   "Carrier_40_G120DStatusWord.3" AT %I2362.3 : Bool;   // Bit_03_FAULT
   "Carrier_40_G120DStatusWord.4" AT %I2362.4 : Bool;   // Bit_04_OFF2
   "Carrier_40_G120DStatusWord.5" AT %I2362.5 : Bool;   // Bit_05_OFF3
   "Carrier_40_G120DStatusWord.6" AT %I2362.6 : Bool;   // Bit_06_LOCK_OUT
   "Carrier_40_G120DStatusWord.7" AT %I2362.7 : Bool;   // Bit_07_WARN
   "Carrier_40_G120DStatusWord.8" AT %I2363.0 : Bool;   // Bit_08_NO_DEVIATION
   "Carrier_40_G120DStatusWord.9" AT %I2363.1 : Bool;   // Bit_09_CONTR_PLC
   "Carrier_40_G120DStatusWord.10" AT %I2363.2 : Bool;   // Bit_10_F_MAX
   "Carrier_40_G120DStatusWord.11" AT %I2363.3 : Bool;   // Bit_11_LIMIT_REACHED
   "Carrier_40_G120DStatusWord.12" AT %I2363.4 : Bool;   // Bit_12_BRAKE_OPEN
   "Carrier_40_G120DStatusWord.13" AT %I2363.5 : Bool;   // Bit_13_NO_OVERTEMP
   "Carrier_40_G120DStatusWord.14" AT %I2363.6 : Bool;   // Bit_14_CW_CCW
   "Carrier_40_G120DStatusWord.15" AT %I2363.7 : Bool;   // Bit_15_OVERL
   "Carrier_40_Slot2_Input" AT %IW2364 : Word;   // SLOT 2 INPUT WORD
   "Carrier_40_CrashDetectSW" AT %I2364.0 : Bool;   // CRASH DETECT SW
   "Carrier_40_SpareSafetyInput(2_1)" AT %I2364.1 : Bool;   // SPARE SAFETY INPUT
   "Carrier_40_SpareSafetyInput(2_2)" AT %I2364.2 : Bool;   // SPARE SAFETY INPUT
   "Carrier_40_SpareSafetyInput(2_3)" AT %I2364.3 : Bool;   // SPARE SAFETY INPUT
   "Carrier_40_SpareSafetyInput(2_4)" AT %I2364.4 : Bool;   // SPARE SAFETY INPUT
   "Carrier_40_SpareSafetyInput(2_5)" AT %I2364.5 : Bool;   // SPARE SAFETY INPUT
   "Carrier_40_SpareSafetyInput(2_6)" AT %I2364.6 : Bool;   // SPARE SAFETY INPUT
   "Carrier_40_SpareSafetyInput(2_7)" AT %I2364.7 : Bool;   // SPARE SAFETY INPUT
   "Carrier_40_Slot3_SafetyOutput" AT %IW2365 : Word;   // SLOT 3 SAFETY OUTPUT WORD
   "Carrier_40_Crash_Detect_OK" AT %I2365.0 : Bool;   // CARRIER CRASH DETECT
   "Carrier_40_SpareSafetyOutput(3_1)" AT %I2365.1 : Bool;   // SPARE SAFETY OUTPUT
   "Carrier_40_SpareSafetyOutput(3_2)" AT %I2365.2 : Bool;   // SPARE SAFETY OUTPUT
   "Carrier_40_SpareSafetyOutput(3_3)" AT %I2365.3 : Bool;   // SPARE SAFETY OUTPUT
   "Carrier_40_SpareSafetyOutput(3_4)" AT %I2365.4 : Bool;   // SPARE SAFETY OUTPUT
   "Carrier_40_SpareSafetyOutput(3_5)" AT %I2365.5 : Bool;   // SPARE SAFETY OUTPUT
   "Carrier_40_SpareSafetyOutput(3_6)" AT %I2365.6 : Bool;   // SPARE SAFETY OUTPUT
   "Carrier_40_SpareSafetyOutput(3_7)" AT %I2365.7 : Bool;   // SPARE SAFETY OUTPUT
   "Carrier_40_Slot4_Input" AT %IW2366 : Word;   // SLOT 4 INPUT WORD
   "Carrier_40_480VPowerOn_MDCB1" AT %I2366.0 : Bool;   // 480 VAC POWER ON MDCB 1
   "Carrier_40_SpareInput(4_1)" AT %I2366.1 : Bool;   // SPARE INPUT
   "Carrier_40_SpareInput(4_2)" AT %I2366.2 : Bool;   // SPARE INPUT
   "Carrier_40_SitopSelectStatus" AT %I2366.3 : Bool;   // SITOP SELECT STATUS
   "Carrier_40_DCsupplyOnPSCB2" AT %I2366.4 : Bool;   // DC SUPPLY ON PSCB 2
   "Carrier_40_SpareInput(4_5)" AT %I2366.5 : Bool;   // SPARE INPUT
   "Carrier_40_SpareInput(4_6)" AT %I2366.6 : Bool;   // SPARE INPUT
   "Carrier_40_SpareInput(4_7)" AT %I2366.7 : Bool;   // SPARE INPUT
   "Carrier_40_PB1_ProdHoldLH" AT %I2367.0 : Bool;   // PB 1 PRODUCTION HOLD LH
   "Carrier_40_PB2_ResetLH" AT %I2367.1 : Bool;   // PB 2 RESET LH
   "Carrier_40_PB3_ProdHoldRH" AT %I2367.2 : Bool;   // PB 3 PRODUCTION HOLD RH
   "Carrier_40_PB4_ResetRH" AT %I2367.3 : Bool;   // PB 4 RESET RH
   "Carrier_40_SpareInput(4_14)" AT %I2367.4 : Bool;   // SPARE INPUT
   "Carrier_40_SpareInput(4_15)" AT %I2367.5 : Bool;   // SPARE INPUT
   "Carrier_40_SpareInput(4_16)" AT %I2367.6 : Bool;   // SPARE INPUT
   "Carrier_40_SpareInput(4_17)" AT %I2367.7 : Bool;   // SPARE INPUT
   "Carrier_40_Slot5_Output" AT %IW2368 : Word;   // SLOT 5 OUTPUT WORD
   "Carrier_40_IRD400_HMI_24VDC_ENABLE" AT %I2368.0 : Bool;   // IRD 400 PANEL HMI 24V DC POWER
   "Carrier_40_FaultLight_LH" AT %I2368.1 : Bool;   // FAULT LIGHT LH
   "Carrier_40_RunLight_LH" AT %I2368.2 : Bool;   // RUN LIGHT LH
   "Carrier_40_FaultLight_RH" AT %I2368.3 : Bool;   // FAULT LIGHT RH
   "Carrier_40_RunLight_RH" AT %I2368.4 : Bool;   // RUN LIGHT RH
   "Carrier_40_SpareOutput(5_5)" AT %I2368.5 : Bool;   // SPARE OUTPUT
   "Carrier_40_SpareOutput(5_6)" AT %I2368.6 : Bool;   // SPARE OUTPUT
   "Carrier_40_SpareOutput(5_7)" AT %I2368.7 : Bool;   // SPARE OUTPUT
   "Carrier_40_ActualSpeed" AT %IW2370 : Word;   // ACTUAL SPEED
   "Carrier_40_CarrierDriveAlarm" AT %IW2372 : Word;   // CARRIER DRIVE ALARM
   "Carrier_40_CarrierDriveWarning" AT %IW2374 : Word;   // CARRIER DRIVE WARNING
   "Carrier_41_Status" AT %IW2400 : Word;   // CARRIER STATUS WORD
   "Carrier_41_Status.0" AT %I2400.0 : Bool;   // HEARTBEAT
   "Carrier_41_Status.1" AT %I2400.1 : Bool;   // MANUAL
   "Carrier_41_Status.2" AT %I2400.2 : Bool;   // IN_AUTO
   "Carrier_41_Status.3" AT %I2400.3 : Bool;   // POSITIONING_COMPLETE
   "Carrier_41_Status.4" AT %I2400.4 : Bool;   // PRODUCTION HOLD
   "Carrier_41_Status.5" AT %I2400.5 : Bool;   // CARRIER MOVING FORWARD
   "Carrier_41_Status.6" AT %I2400.6 : Bool;   // CARRIER MOVING REVERSE
   "Carrier_41_Status.7" AT %I2400.7 : Bool;   // CARRIER FAULT
   "Carrier_41_Status.8" AT %I2401.0 : Bool;   // CRASH DETECT TRIPPED
   "Carrier_41_Status.9" AT %I2401.1 : Bool;
   "Carrier_41_Status.10" AT %I2401.2 : Bool;
   "Carrier_41_Status.11" AT %I2401.3 : Bool;
   "Carrier_41_Status.12" AT %I2401.4 : Bool;
   "Carrier_41_Status.13" AT %I2401.5 : Bool;
   "Carrier_41_Status.14" AT %I2401.6 : Bool;
   "Carrier_41_Status.15" AT %I2401.7 : Bool;
   "Carrier_41_SDCFaultCode" AT %IW2402 : Word;   // SDC FAULT CODE
   "Carrier_41_CarrierPosition" AT %ID2404 : DWord;   // CARRIER POSITION
   "Carrier_41_CarrierNumber" AT %IW2408 : Word;   // CARRIER NUMBER
   "Carrier_41_G120DControlWord" AT %IW2410 : Word;   // G120D_STW1_CONTROL
   "Carrier_41_G120DControlWord.0" AT %I2410.0 : Bool;   // Bit_00_ON
   "Carrier_41_G120DControlWord.1" AT %I2410.1 : Bool;   // Bit_01_AUS2_INH
   "Carrier_41_G120DControlWord.2" AT %I2410.2 : Bool;   // Bit_02_AUS3_STOP
   "Carrier_41_G120DControlWord.3" AT %I2410.3 : Bool;   // Bit_03_EN
   "Carrier_41_G120DControlWord.4" AT %I2410.4 : Bool;   // Bit_04_EN_RAMP
   "Carrier_41_G120DControlWord.5" AT %I2410.5 : Bool;   // Bit_05_START_RAMP
   "Carrier_41_G120DControlWord.6" AT %I2410.6 : Bool;   // Bit_06_SETPOINT
   "Carrier_41_G120DControlWord.7" AT %I2410.7 : Bool;   // Bit_07_RESET
   "Carrier_41_G120DControlWord.8" AT %I2411.0 : Bool;   // Bit_08_JOG_R
   "Carrier_41_G120DControlWord.9" AT %I2411.1 : Bool;   // Bit_09_JOG_L
   "Carrier_41_G120DControlWord.10" AT %I2411.2 : Bool;   // Bit_10_CONTR_PLC
   "Carrier_41_G120DControlWord.11" AT %I2411.3 : Bool;   // Bit_11_REVERSE
   "Carrier_41_G120DControlWord.12" AT %I2411.4 : Bool;   // Bit_12_BRAKE_RELEASE
   "Carrier_41_G120DControlWord.13" AT %I2411.5 : Bool;   // Bit_13_DDS
   "Carrier_41_G120DControlWord.14" AT %I2411.6 : Bool;   // Bit_14_DO0
   "Carrier_41_G120DControlWord.15" AT %I2411.7 : Bool;   // Bit_15_DO1
   "Carrier_41_G120DStatusWord" AT %IW2412 : Word;   // G120D_ZSW1_STATUS
   "Carrier_41_G120DStatusWord.0" AT %I2412.0 : Bool;   // Bit_00_READY_RUN
   "Carrier_41_G120DStatusWord.1" AT %I2412.1 : Bool;   // Bit_01_READY_ON
   "Carrier_41_G120DStatusWord.2" AT %I2412.2 : Bool;   // Bit_02_ENABLE
   "Carrier_41_G120DStatusWord.3" AT %I2412.3 : Bool;   // Bit_03_FAULT
   "Carrier_41_G120DStatusWord.4" AT %I2412.4 : Bool;   // Bit_04_OFF2
   "Carrier_41_G120DStatusWord.5" AT %I2412.5 : Bool;   // Bit_05_OFF3
   "Carrier_41_G120DStatusWord.6" AT %I2412.6 : Bool;   // Bit_06_LOCK_OUT
   "Carrier_41_G120DStatusWord.7" AT %I2412.7 : Bool;   // Bit_07_WARN
   "Carrier_41_G120DStatusWord.8" AT %I2413.0 : Bool;   // Bit_08_NO_DEVIATION
   "Carrier_41_G120DStatusWord.9" AT %I2413.1 : Bool;   // Bit_09_CONTR_PLC
   "Carrier_41_G120DStatusWord.10" AT %I2413.2 : Bool;   // Bit_10_F_MAX
   "Carrier_41_G120DStatusWord.11" AT %I2413.3 : Bool;   // Bit_11_LIMIT_REACHED
   "Carrier_41_G120DStatusWord.12" AT %I2413.4 : Bool;   // Bit_12_BRAKE_OPEN
   "Carrier_41_G120DStatusWord.13" AT %I2413.5 : Bool;   // Bit_13_NO_OVERTEMP
   "Carrier_41_G120DStatusWord.14" AT %I2413.6 : Bool;   // Bit_14_CW_CCW
   "Carrier_41_G120DStatusWord.15" AT %I2413.7 : Bool;   // Bit_15_OVERL
   "Carrier_41_Slot2_Input" AT %IW2414 : Word;   // SLOT 2 INPUT WORD
   "Carrier_41_CrashDetectSW" AT %I2414.0 : Bool;   // CRASH DETECT SW
   "Carrier_41_SpareSafetyInput(2_1)" AT %I2414.1 : Bool;   // SPARE SAFETY INPUT
   "Carrier_41_SpareSafetyInput(2_2)" AT %I2414.2 : Bool;   // SPARE SAFETY INPUT
   "Carrier_41_SpareSafetyInput(2_3)" AT %I2414.3 : Bool;   // SPARE SAFETY INPUT
   "Carrier_41_SpareSafetyInput(2_4)" AT %I2414.4 : Bool;   // SPARE SAFETY INPUT
   "Carrier_41_SpareSafetyInput(2_5)" AT %I2414.5 : Bool;   // SPARE SAFETY INPUT
   "Carrier_41_SpareSafetyInput(2_6)" AT %I2414.6 : Bool;   // SPARE SAFETY INPUT
   "Carrier_41_SpareSafetyInput(2_7)" AT %I2414.7 : Bool;   // SPARE SAFETY INPUT
   "Carrier_41_Slot3_SafetyOutput" AT %IW2415 : Word;   // SLOT 3 SAFETY OUTPUT WORD
   "Carrier_41_Crash_Detect_OK" AT %I2415.0 : Bool;   // CARRIER CRASH DETECT
   "Carrier_41_SpareSafetyOutput(3_1)" AT %I2415.1 : Bool;   // SPARE SAFETY OUTPUT
   "Carrier_41_SpareSafetyOutput(3_2)" AT %I2415.2 : Bool;   // SPARE SAFETY OUTPUT
   "Carrier_41_SpareSafetyOutput(3_3)" AT %I2415.3 : Bool;   // SPARE SAFETY OUTPUT
   "Carrier_41_SpareSafetyOutput(3_4)" AT %I2415.4 : Bool;   // SPARE SAFETY OUTPUT
   "Carrier_41_SpareSafetyOutput(3_5)" AT %I2415.5 : Bool;   // SPARE SAFETY OUTPUT
   "Carrier_41_SpareSafetyOutput(3_6)" AT %I2415.6 : Bool;   // SPARE SAFETY OUTPUT
   "Carrier_41_SpareSafetyOutput(3_7)" AT %I2415.7 : Bool;   // SPARE SAFETY OUTPUT
   "Carrier_41_Slot4_Input" AT %IW2416 : Word;   // SLOT 4 INPUT WORD
   "Carrier_41_480VPowerOn_MDCB1" AT %I2416.0 : Bool;   // 480 VAC POWER ON MDCB 1
   "Carrier_41_SpareInput(4_1)" AT %I2416.1 : Bool;   // SPARE INPUT
   "Carrier_41_SpareInput(4_2)" AT %I2416.2 : Bool;   // SPARE INPUT
   "Carrier_41_SitopSelectStatus" AT %I2416.3 : Bool;   // SITOP SELECT STATUS
   "Carrier_41_DCsupplyOnPSCB2" AT %I2416.4 : Bool;   // DC SUPPLY ON PSCB 2
   "Carrier_41_SpareInput(4_5)" AT %I2416.5 : Bool;   // SPARE INPUT
   "Carrier_41_SpareInput(4_6)" AT %I2416.6 : Bool;   // SPARE INPUT
   "Carrier_41_SpareInput(4_7)" AT %I2416.7 : Bool;   // SPARE INPUT
   "Carrier_41_PB1_ProdHoldLH" AT %I2417.0 : Bool;   // PB 1 PRODUCTION HOLD LH
   "Carrier_41_PB2_ResetLH" AT %I2417.1 : Bool;   // PB 2 RESET LH
   "Carrier_41_PB3_ProdHoldRH" AT %I2417.2 : Bool;   // PB 3 PRODUCTION HOLD RH
   "Carrier_41_PB4_ResetRH" AT %I2417.3 : Bool;   // PB 4 RESET RH
   "Carrier_41_SpareInput(4_14)" AT %I2417.4 : Bool;   // SPARE INPUT
   "Carrier_41_SpareInput(4_15)" AT %I2417.5 : Bool;   // SPARE INPUT
   "Carrier_41_SpareInput(4_16)" AT %I2417.6 : Bool;   // SPARE INPUT
   "Carrier_41_SpareInput(4_17)" AT %I2417.7 : Bool;   // SPARE INPUT
   "Carrier_41_Slot5_Output" AT %IW2418 : Word;   // SLOT 5 OUTPUT WORD
   "Carrier_41_IRD400_HMI_24VDC_ENABLE" AT %I2418.0 : Bool;   // IRD 400 PANEL HMI 24V DC POWER
   "Carrier_41_FaultLight_LH" AT %I2418.1 : Bool;   // FAULT LIGHT LH
   "Carrier_41_RunLight_LH" AT %I2418.2 : Bool;   // RUN LIGHT LH
   "Carrier_41_FaultLight_RH" AT %I2418.3 : Bool;   // FAULT LIGHT RH
   "Carrier_41_RunLight_RH" AT %I2418.4 : Bool;   // RUN LIGHT RH
   "Carrier_41_SpareOutput(5_5)" AT %I2418.5 : Bool;   // SPARE OUTPUT
   "Carrier_41_SpareOutput(5_6)" AT %I2418.6 : Bool;   // SPARE OUTPUT
   "Carrier_41_SpareOutput(5_7)" AT %I2418.7 : Bool;   // SPARE OUTPUT
   "Carrier_41_ActualSpeed" AT %IW2420 : Word;   // ACTUAL SPEED
   "Carrier_41_CarrierDriveAlarm" AT %IW2422 : Word;   // CARRIER DRIVE ALARM
   "Carrier_41_CarrierDriveWarning" AT %IW2424 : Word;   // CARRIER DRIVE WARNING
   "Carrier_42_Status" AT %IW2450 : Word;   // CARRIER STATUS WORD
   "Carrier_42_Status.0" AT %I2450.0 : Bool;   // HEARTBEAT
   "Carrier_42_Status.1" AT %I2450.1 : Bool;   // MANUAL
   "Carrier_42_Status.2" AT %I2450.2 : Bool;   // IN_AUTO
   "Carrier_42_Status.3" AT %I2450.3 : Bool;   // POSITIONING_COMPLETE
   "Carrier_42_Status.4" AT %I2450.4 : Bool;   // PRODUCTION HOLD
   "Carrier_42_Status.5" AT %I2450.5 : Bool;   // CARRIER MOVING FORWARD
   "Carrier_42_Status.6" AT %I2450.6 : Bool;   // CARRIER MOVING REVERSE
   "Carrier_42_Status.7" AT %I2450.7 : Bool;   // CARRIER FAULT
   "Carrier_42_Status.8" AT %I2451.0 : Bool;   // CRASH DETECT TRIPPED
   "Carrier_42_Status.9" AT %I2451.1 : Bool;
   "Carrier_42_Status.10" AT %I2451.2 : Bool;
   "Carrier_42_Status.11" AT %I2451.3 : Bool;
   "Carrier_42_Status.12" AT %I2451.4 : Bool;
   "Carrier_42_Status.13" AT %I2451.5 : Bool;
   "Carrier_42_Status.14" AT %I2451.6 : Bool;
   "Carrier_42_Status.15" AT %I2451.7 : Bool;
   "Carrier_42_SDCFaultCode" AT %IW2452 : Word;   // SDC FAULT CODE
   "Carrier_42_CarrierPosition" AT %ID2454 : DWord;   // CARRIER POSITION
   "Carrier_42_CarrierNumber" AT %IW2458 : Word;   // CARRIER NUMBER
   "Carrier_42_G120DControlWord" AT %IW2460 : Word;   // G120D_STW1_CONTROL
   "Carrier_42_G120DControlWord.0" AT %I2460.0 : Bool;   // Bit_00_ON
   "Carrier_42_G120DControlWord.1" AT %I2460.1 : Bool;   // Bit_01_AUS2_INH
   "Carrier_42_G120DControlWord.2" AT %I2460.2 : Bool;   // Bit_02_AUS3_STOP
   "Carrier_42_G120DControlWord.3" AT %I2460.3 : Bool;   // Bit_03_EN
   "Carrier_42_G120DControlWord.4" AT %I2460.4 : Bool;   // Bit_04_EN_RAMP
   "Carrier_42_G120DControlWord.5" AT %I2460.5 : Bool;   // Bit_05_START_RAMP
   "Carrier_42_G120DControlWord.6" AT %I2460.6 : Bool;   // Bit_06_SETPOINT
   "Carrier_42_G120DControlWord.7" AT %I2460.7 : Bool;   // Bit_07_RESET
   "Carrier_42_G120DControlWord.8" AT %I2461.0 : Bool;   // Bit_08_JOG_R
   "Carrier_42_G120DControlWord.9" AT %I2461.1 : Bool;   // Bit_09_JOG_L
   "Carrier_42_G120DControlWord.10" AT %I2461.2 : Bool;   // Bit_10_CONTR_PLC
   "Carrier_42_G120DControlWord.11" AT %I2461.3 : Bool;   // Bit_11_REVERSE
   "Carrier_42_G120DControlWord.12" AT %I2461.4 : Bool;   // Bit_12_BRAKE_RELEASE
   "Carrier_42_G120DControlWord.13" AT %I2461.5 : Bool;   // Bit_13_DDS
   "Carrier_42_G120DControlWord.14" AT %I2461.6 : Bool;   // Bit_14_DO0
   "Carrier_42_G120DControlWord.15" AT %I2461.7 : Bool;   // Bit_15_DO1
   "Carrier_42_G120DStatusWord" AT %IW2462 : Word;   // G120D_ZSW1_STATUS
   "Carrier_42_G120DStatusWord.0" AT %I2462.0 : Bool;   // Bit_00_READY_RUN
   "Carrier_42_G120DStatusWord.1" AT %I2462.1 : Bool;   // Bit_01_READY_ON
   "Carrier_42_G120DStatusWord.2" AT %I2462.2 : Bool;   // Bit_02_ENABLE
   "Carrier_42_G120DStatusWord.3" AT %I2462.3 : Bool;   // Bit_03_FAULT
   "Carrier_42_G120DStatusWord.4" AT %I2462.4 : Bool;   // Bit_04_OFF2
   "Carrier_42_G120DStatusWord.5" AT %I2462.5 : Bool;   // Bit_05_OFF3
   "Carrier_42_G120DStatusWord.6" AT %I2462.6 : Bool;   // Bit_06_LOCK_OUT
   "Carrier_42_G120DStatusWord.7" AT %I2462.7 : Bool;   // Bit_07_WARN
   "Carrier_42_G120DStatusWord.8" AT %I2463.0 : Bool;   // Bit_08_NO_DEVIATION
   "Carrier_42_G120DStatusWord.9" AT %I2463.1 : Bool;   // Bit_09_CONTR_PLC
   "Carrier_42_G120DStatusWord.10" AT %I2463.2 : Bool;   // Bit_10_F_MAX
   "Carrier_42_G120DStatusWord.11" AT %I2463.3 : Bool;   // Bit_11_LIMIT_REACHED
   "Carrier_42_G120DStatusWord.12" AT %I2463.4 : Bool;   // Bit_12_BRAKE_OPEN
   "Carrier_42_G120DStatusWord.13" AT %I2463.5 : Bool;   // Bit_13_NO_OVERTEMP
   "Carrier_42_G120DStatusWord.14" AT %I2463.6 : Bool;   // Bit_14_CW_CCW
   "Carrier_42_G120DStatusWord.15" AT %I2463.7 : Bool;   // Bit_15_OVERL
   "Carrier_42_Slot2_Input" AT %IW2464 : Word;   // SLOT 2 INPUT WORD
   "Carrier_42_CrashDetectSW" AT %I2464.0 : Bool;   // CRASH DETECT SW
   "Carrier_42_SpareSafetyInput(2_1)" AT %I2464.1 : Bool;   // SPARE SAFETY INPUT
   "Carrier_42_SpareSafetyInput(2_2)" AT %I2464.2 : Bool;   // SPARE SAFETY INPUT
   "Carrier_42_SpareSafetyInput(2_3)" AT %I2464.3 : Bool;   // SPARE SAFETY INPUT
   "Carrier_42_SpareSafetyInput(2_4)" AT %I2464.4 : Bool;   // SPARE SAFETY INPUT
   "Carrier_42_SpareSafetyInput(2_5)" AT %I2464.5 : Bool;   // SPARE SAFETY INPUT
   "Carrier_42_SpareSafetyInput(2_6)" AT %I2464.6 : Bool;   // SPARE SAFETY INPUT
   "Carrier_42_SpareSafetyInput(2_7)" AT %I2464.7 : Bool;   // SPARE SAFETY INPUT
   "Carrier_42_Slot3_SafetyOutput" AT %IW2465 : Word;   // SLOT 3 SAFETY OUTPUT WORD
   "Carrier_42_Crash_Detect_OK" AT %I2465.0 : Bool;   // CARRIER CRASH DETECT
   "Carrier_42_SpareSafetyOutput(3_1)" AT %I2465.1 : Bool;   // SPARE SAFETY OUTPUT
   "Carrier_42_SpareSafetyOutput(3_2)" AT %I2465.2 : Bool;   // SPARE SAFETY OUTPUT
   "Carrier_42_SpareSafetyOutput(3_3)" AT %I2465.3 : Bool;   // SPARE SAFETY OUTPUT
   "Carrier_42_SpareSafetyOutput(3_4)" AT %I2465.4 : Bool;   // SPARE SAFETY OUTPUT
   "Carrier_42_SpareSafetyOutput(3_5)" AT %I2465.5 : Bool;   // SPARE SAFETY OUTPUT
   "Carrier_42_SpareSafetyOutput(3_6)" AT %I2465.6 : Bool;   // SPARE SAFETY OUTPUT
   "Carrier_42_SpareSafetyOutput(3_7)" AT %I2465.7 : Bool;   // SPARE SAFETY OUTPUT
   "Carrier_42_Slot4_Input" AT %IW2466 : Word;   // SLOT 4 INPUT WORD
   "Carrier_42_480VPowerOn_MDCB1" AT %I2466.0 : Bool;   // 480 VAC POWER ON MDCB 1
   "Carrier_42_SpareInput(4_1)" AT %I2466.1 : Bool;   // SPARE INPUT
   "Carrier_42_SpareInput(4_2)" AT %I2466.2 : Bool;   // SPARE INPUT
   "Carrier_42_SitopSelectStatus" AT %I2466.3 : Bool;   // SITOP SELECT STATUS
   "Carrier_42_DCsupplyOnPSCB2" AT %I2466.4 : Bool;   // DC SUPPLY ON PSCB 2
   "Carrier_42_SpareInput(4_5)" AT %I2466.5 : Bool;   // SPARE INPUT
   "Carrier_42_SpareInput(4_6)" AT %I2466.6 : Bool;   // SPARE INPUT
   "Carrier_42_SpareInput(4_7)" AT %I2466.7 : Bool;   // SPARE INPUT
   "Carrier_42_PB1_ProdHoldLH" AT %I2467.0 : Bool;   // PB 1 PRODUCTION HOLD LH
   "Carrier_42_PB2_ResetLH" AT %I2467.1 : Bool;   // PB 2 RESET LH
   "Carrier_42_PB3_ProdHoldRH" AT %I2467.2 : Bool;   // PB 3 PRODUCTION HOLD RH
   "Carrier_42_PB4_ResetRH" AT %I2467.3 : Bool;   // PB 4 RESET RH
   "Carrier_42_SpareInput(4_14)" AT %I2467.4 : Bool;   // SPARE INPUT
   "Carrier_42_SpareInput(4_15)" AT %I2467.5 : Bool;   // SPARE INPUT
   "Carrier_42_SpareInput(4_16)" AT %I2467.6 : Bool;   // SPARE INPUT
   "Carrier_42_SpareInput(4_17)" AT %I2467.7 : Bool;   // SPARE INPUT
   "Carrier_42_Slot5_Output" AT %IW2468 : Word;   // SLOT 5 OUTPUT WORD
   "Carrier_42_IRD400_HMI_24VDC_ENABLE" AT %I2468.0 : Bool;   // IRD 400 PANEL HMI 24V DC POWER
   "Carrier_42_FaultLight_LH" AT %I2468.1 : Bool;   // FAULT LIGHT LH
   "Carrier_42_RunLight_LH" AT %I2468.2 : Bool;   // RUN LIGHT LH
   "Carrier_42_FaultLight_RH" AT %I2468.3 : Bool;   // FAULT LIGHT RH
   "Carrier_42_RunLight_RH" AT %I2468.4 : Bool;   // RUN LIGHT RH
   "Carrier_42_SpareOutput(5_5)" AT %I2468.5 : Bool;   // SPARE OUTPUT
   "Carrier_42_SpareOutput(5_6)" AT %I2468.6 : Bool;   // SPARE OUTPUT
   "Carrier_42_SpareOutput(5_7)" AT %I2468.7 : Bool;   // SPARE OUTPUT
   "Carrier_42_ActualSpeed" AT %IW2470 : Word;   // ACTUAL SPEED
   "Carrier_42_CarrierDriveAlarm" AT %IW2472 : Word;   // CARRIER DRIVE ALARM
   "Carrier_42_CarrierDriveWarning" AT %IW2474 : Word;   // CARRIER DRIVE WARNING
   "Carrier_43_Status" AT %IW2500 : Word;   // CARRIER STATUS WORD
   "Carrier_43_Status.0" AT %I2500.0 : Bool;   // HEARTBEAT
   "Carrier_43_Status.1" AT %I2500.1 : Bool;   // MANUAL
   "Carrier_43_Status.2" AT %I2500.2 : Bool;   // IN_AUTO
   "Carrier_43_Status.3" AT %I2500.3 : Bool;   // POSITIONING_COMPLETE
   "Carrier_43_Status.4" AT %I2500.4 : Bool;   // PRODUCTION HOLD
   "Carrier_43_Status.5" AT %I2500.5 : Bool;   // CARRIER MOVING FORWARD
   "Carrier_43_Status.6" AT %I2500.6 : Bool;   // CARRIER MOVING REVERSE
   "Carrier_43_Status.7" AT %I2500.7 : Bool;   // CARRIER FAULT
   "Carrier_43_Status.8" AT %I2501.0 : Bool;   // CRASH DETECT TRIPPED
   "Carrier_43_Status.9" AT %I2501.1 : Bool;
   "Carrier_43_Status.10" AT %I2501.2 : Bool;
   "Carrier_43_Status.11" AT %I2501.3 : Bool;
   "Carrier_43_Status.12" AT %I2501.4 : Bool;
   "Carrier_43_Status.13" AT %I2501.5 : Bool;
   "Carrier_43_Status.14" AT %I2501.6 : Bool;
   "Carrier_43_Status.15" AT %I2501.7 : Bool;
   "Carrier_43_SDCFaultCode" AT %IW2502 : Word;   // SDC FAULT CODE
   "Carrier_43_CarrierPosition" AT %ID2504 : DWord;   // CARRIER POSITION
   "Carrier_43_CarrierNumber" AT %IW2508 : Word;   // CARRIER NUMBER
   "Carrier_43_G120DControlWord" AT %IW2510 : Word;   // G120D_STW1_CONTROL
   "Carrier_43_G120DControlWord.0" AT %I2510.0 : Bool;   // Bit_00_ON
   "Carrier_43_G120DControlWord.1" AT %I2510.1 : Bool;   // Bit_01_AUS2_INH
   "Carrier_43_G120DControlWord.2" AT %I2510.2 : Bool;   // Bit_02_AUS3_STOP
   "Carrier_43_G120DControlWord.3" AT %I2510.3 : Bool;   // Bit_03_EN
   "Carrier_43_G120DControlWord.4" AT %I2510.4 : Bool;   // Bit_04_EN_RAMP
   "Carrier_43_G120DControlWord.5" AT %I2510.5 : Bool;   // Bit_05_START_RAMP
   "Carrier_43_G120DControlWord.6" AT %I2510.6 : Bool;   // Bit_06_SETPOINT
   "Carrier_43_G120DControlWord.7" AT %I2510.7 : Bool;   // Bit_07_RESET
   "Carrier_43_G120DControlWord.8" AT %I2511.0 : Bool;   // Bit_08_JOG_R
   "Carrier_43_G120DControlWord.9" AT %I2511.1 : Bool;   // Bit_09_JOG_L
   "Carrier_43_G120DControlWord.10" AT %I2511.2 : Bool;   // Bit_10_CONTR_PLC
   "Carrier_43_G120DControlWord.11" AT %I2511.3 : Bool;   // Bit_11_REVERSE
   "Carrier_43_G120DControlWord.12" AT %I2511.4 : Bool;   // Bit_12_BRAKE_RELEASE
   "Carrier_43_G120DControlWord.13" AT %I2511.5 : Bool;   // Bit_13_DDS
   "Carrier_43_G120DControlWord.14" AT %I2511.6 : Bool;   // Bit_14_DO0
   "Carrier_43_G120DControlWord.15" AT %I2511.7 : Bool;   // Bit_15_DO1
   "Carrier_43_G120DStatusWord" AT %IW2512 : Word;   // G120D_ZSW1_STATUS
   "Carrier_43_G120DStatusWord.0" AT %I2512.0 : Bool;   // Bit_00_READY_RUN
   "Carrier_43_G120DStatusWord.1" AT %I2512.1 : Bool;   // Bit_01_READY_ON
   "Carrier_43_G120DStatusWord.2" AT %I2512.2 : Bool;   // Bit_02_ENABLE
   "Carrier_43_G120DStatusWord.3" AT %I2512.3 : Bool;   // Bit_03_FAULT
   "Carrier_43_G120DStatusWord.4" AT %I2512.4 : Bool;   // Bit_04_OFF2
   "Carrier_43_G120DStatusWord.5" AT %I2512.5 : Bool;   // Bit_05_OFF3
   "Carrier_43_G120DStatusWord.6" AT %I2512.6 : Bool;   // Bit_06_LOCK_OUT
   "Carrier_43_G120DStatusWord.7" AT %I2512.7 : Bool;   // Bit_07_WARN
   "Carrier_43_G120DStatusWord.8" AT %I2513.0 : Bool;   // Bit_08_NO_DEVIATION
   "Carrier_43_G120DStatusWord.9" AT %I2513.1 : Bool;   // Bit_09_CONTR_PLC
   "Carrier_43_G120DStatusWord.10" AT %I2513.2 : Bool;   // Bit_10_F_MAX
   "Carrier_43_G120DStatusWord.11" AT %I2513.3 : Bool;   // Bit_11_LIMIT_REACHED
   "Carrier_43_G120DStatusWord.12" AT %I2513.4 : Bool;   // Bit_12_BRAKE_OPEN
   "Carrier_43_G120DStatusWord.13" AT %I2513.5 : Bool;   // Bit_13_NO_OVERTEMP
   "Carrier_43_G120DStatusWord.14" AT %I2513.6 : Bool;   // Bit_14_CW_CCW
   "Carrier_43_G120DStatusWord.15" AT %I2513.7 : Bool;   // Bit_15_OVERL
   "Carrier_43_Slot2_Input" AT %IW2514 : Word;   // SLOT 2 INPUT WORD
   "Carrier_43_CrashDetectSW" AT %I2514.0 : Bool;   // CRASH DETECT SW
   "Carrier_43_SpareSafetyInput(2_1)" AT %I2514.1 : Bool;   // SPARE SAFETY INPUT
   "Carrier_43_SpareSafetyInput(2_2)" AT %I2514.2 : Bool;   // SPARE SAFETY INPUT
   "Carrier_43_SpareSafetyInput(2_3)" AT %I2514.3 : Bool;   // SPARE SAFETY INPUT
   "Carrier_43_SpareSafetyInput(2_4)" AT %I2514.4 : Bool;   // SPARE SAFETY INPUT
   "Carrier_43_SpareSafetyInput(2_5)" AT %I2514.5 : Bool;   // SPARE SAFETY INPUT
   "Carrier_43_SpareSafetyInput(2_6)" AT %I2514.6 : Bool;   // SPARE SAFETY INPUT
   "Carrier_43_SpareSafetyInput(2_7)" AT %I2514.7 : Bool;   // SPARE SAFETY INPUT
   "Carrier_43_Slot3_SafetyOutput" AT %IW2515 : Word;   // SLOT 3 SAFETY OUTPUT WORD
   "Carrier_43_Crash_Detect_OK" AT %I2515.0 : Bool;   // CARRIER CRASH DETECT
   "Carrier_43_SpareSafetyOutput(3_1)" AT %I2515.1 : Bool;   // SPARE SAFETY OUTPUT
   "Carrier_43_SpareSafetyOutput(3_2)" AT %I2515.2 : Bool;   // SPARE SAFETY OUTPUT
   "Carrier_43_SpareSafetyOutput(3_3)" AT %I2515.3 : Bool;   // SPARE SAFETY OUTPUT
   "Carrier_43_SpareSafetyOutput(3_4)" AT %I2515.4 : Bool;   // SPARE SAFETY OUTPUT
   "Carrier_43_SpareSafetyOutput(3_5)" AT %I2515.5 : Bool;   // SPARE SAFETY OUTPUT
   "Carrier_43_SpareSafetyOutput(3_6)" AT %I2515.6 : Bool;   // SPARE SAFETY OUTPUT
   "Carrier_43_SpareSafetyOutput(3_7)" AT %I2515.7 : Bool;   // SPARE SAFETY OUTPUT
   "Carrier_43_Slot4_Input" AT %IW2516 : Word;   // SLOT 4 INPUT WORD
   "Carrier_43_480VPowerOn_MDCB1" AT %I2516.0 : Bool;   // 480 VAC POWER ON MDCB 1
   "Carrier_43_SpareInput(4_1)" AT %I2516.1 : Bool;   // SPARE INPUT
   "Carrier_43_SpareInput(4_2)" AT %I2516.2 : Bool;   // SPARE INPUT
   "Carrier_43_SitopSelectStatus" AT %I2516.3 : Bool;   // SITOP SELECT STATUS
   "Carrier_43_DCsupplyOnPSCB2" AT %I2516.4 : Bool;   // DC SUPPLY ON PSCB 2
   "Carrier_43_SpareInput(4_5)" AT %I2516.5 : Bool;   // SPARE INPUT
   "Carrier_43_SpareInput(4_6)" AT %I2516.6 : Bool;   // SPARE INPUT
   "Carrier_43_SpareInput(4_7)" AT %I2516.7 : Bool;   // SPARE INPUT
   "Carrier_43_PB1_ProdHoldLH" AT %I2517.0 : Bool;   // PB 1 PRODUCTION HOLD LH
   "Carrier_43_PB2_ResetLH" AT %I2517.1 : Bool;   // PB 2 RESET LH
   "Carrier_43_PB3_ProdHoldRH" AT %I2517.2 : Bool;   // PB 3 PRODUCTION HOLD RH
   "Carrier_43_PB4_ResetRH" AT %I2517.3 : Bool;   // PB 4 RESET RH
   "Carrier_43_SpareInput(4_14)" AT %I2517.4 : Bool;   // SPARE INPUT
   "Carrier_43_SpareInput(4_15)" AT %I2517.5 : Bool;   // SPARE INPUT
   "Carrier_43_SpareInput(4_16)" AT %I2517.6 : Bool;   // SPARE INPUT
   "Carrier_43_SpareInput(4_17)" AT %I2517.7 : Bool;   // SPARE INPUT
   "Carrier_43_Slot5_Output" AT %IW2518 : Word;   // SLOT 5 OUTPUT WORD
   "Carrier_43_IRD400_HMI_24VDC_ENABLE" AT %I2518.0 : Bool;   // IRD 400 PANEL HMI 24V DC POWER
   "Carrier_43_FaultLight_LH" AT %I2518.1 : Bool;   // FAULT LIGHT LH
   "Carrier_43_RunLight_LH" AT %I2518.2 : Bool;   // RUN LIGHT LH
   "Carrier_43_FaultLight_RH" AT %I2518.3 : Bool;   // FAULT LIGHT RH
   "Carrier_43_RunLight_RH" AT %I2518.4 : Bool;   // RUN LIGHT RH
   "Carrier_43_SpareOutput(5_5)" AT %I2518.5 : Bool;   // SPARE OUTPUT
   "Carrier_43_SpareOutput(5_6)" AT %I2518.6 : Bool;   // SPARE OUTPUT
   "Carrier_43_SpareOutput(5_7)" AT %I2518.7 : Bool;   // SPARE OUTPUT
   "Carrier_43_ActualSpeed" AT %IW2520 : Word;   // ACTUAL SPEED
   "Carrier_43_CarrierDriveAlarm" AT %IW2522 : Word;   // CARRIER DRIVE ALARM
   "Carrier_43_CarrierDriveWarning" AT %IW2524 : Word;   // CARRIER DRIVE WARNING
   "Carrier_44_Status" AT %IW2550 : Word;   // CARRIER STATUS WORD
   "Carrier_44_Status.0" AT %I2550.0 : Bool;   // HEARTBEAT
   "Carrier_44_Status.1" AT %I2550.1 : Bool;   // MANUAL
   "Carrier_44_Status.2" AT %I2550.2 : Bool;   // IN_AUTO
   "Carrier_44_Status.3" AT %I2550.3 : Bool;   // POSITIONING_COMPLETE
   "Carrier_44_Status.4" AT %I2550.4 : Bool;   // PRODUCTION HOLD
   "Carrier_44_Status.5" AT %I2550.5 : Bool;   // CARRIER MOVING FORWARD
   "Carrier_44_Status.6" AT %I2550.6 : Bool;   // CARRIER MOVING REVERSE
   "Carrier_44_Status.7" AT %I2550.7 : Bool;   // CARRIER FAULT
   "Carrier_44_Status.8" AT %I2551.0 : Bool;   // CRASH DETECT TRIPPED
   "Carrier_44_Status.9" AT %I2551.1 : Bool;
   "Carrier_44_Status.10" AT %I2551.2 : Bool;
   "Carrier_44_Status.11" AT %I2551.3 : Bool;
   "Carrier_44_Status.12" AT %I2551.4 : Bool;
   "Carrier_44_Status.13" AT %I2551.5 : Bool;
   "Carrier_44_Status.14" AT %I2551.6 : Bool;
   "Carrier_44_Status.15" AT %I2551.7 : Bool;
   "Carrier_44_SDCFaultCode" AT %IW2552 : Word;   // SDC FAULT CODE
   "Carrier_44_CarrierPosition" AT %ID2554 : DWord;   // CARRIER POSITION
   "Carrier_44_CarrierNumber" AT %IW2558 : Word;   // CARRIER NUMBER
   "Carrier_44_G120DControlWord" AT %IW2560 : Word;   // G120D_STW1_CONTROL
   "Carrier_44_G120DControlWord.0" AT %I2560.0 : Bool;   // Bit_00_ON
   "Carrier_44_G120DControlWord.1" AT %I2560.1 : Bool;   // Bit_01_AUS2_INH
   "Carrier_44_G120DControlWord.2" AT %I2560.2 : Bool;   // Bit_02_AUS3_STOP
   "Carrier_44_G120DControlWord.3" AT %I2560.3 : Bool;   // Bit_03_EN
   "Carrier_44_G120DControlWord.4" AT %I2560.4 : Bool;   // Bit_04_EN_RAMP
   "Carrier_44_G120DControlWord.5" AT %I2560.5 : Bool;   // Bit_05_START_RAMP
   "Carrier_44_G120DControlWord.6" AT %I2560.6 : Bool;   // Bit_06_SETPOINT
   "Carrier_44_G120DControlWord.7" AT %I2560.7 : Bool;   // Bit_07_RESET
   "Carrier_44_G120DControlWord.8" AT %I2561.0 : Bool;   // Bit_08_JOG_R
   "Carrier_44_G120DControlWord.9" AT %I2561.1 : Bool;   // Bit_09_JOG_L
   "Carrier_44_G120DControlWord.10" AT %I2561.2 : Bool;   // Bit_10_CONTR_PLC
   "Carrier_44_G120DControlWord.11" AT %I2561.3 : Bool;   // Bit_11_REVERSE
   "Carrier_44_G120DControlWord.12" AT %I2561.4 : Bool;   // Bit_12_BRAKE_RELEASE
   "Carrier_44_G120DControlWord.13" AT %I2561.5 : Bool;   // Bit_13_DDS
   "Carrier_44_G120DControlWord.14" AT %I2561.6 : Bool;   // Bit_14_DO0
   "Carrier_44_G120DControlWord.15" AT %I2561.7 : Bool;   // Bit_15_DO1
   "Carrier_44_G120DStatusWord" AT %IW2562 : Word;   // G120D_ZSW1_STATUS
   "Carrier_44_G120DStatusWord.0" AT %I2562.0 : Bool;   // Bit_00_READY_RUN
   "Carrier_44_G120DStatusWord.1" AT %I2562.1 : Bool;   // Bit_01_READY_ON
   "Carrier_44_G120DStatusWord.2" AT %I2562.2 : Bool;   // Bit_02_ENABLE
   "Carrier_44_G120DStatusWord.3" AT %I2562.3 : Bool;   // Bit_03_FAULT
   "Carrier_44_G120DStatusWord.4" AT %I2562.4 : Bool;   // Bit_04_OFF2
   "Carrier_44_G120DStatusWord.5" AT %I2562.5 : Bool;   // Bit_05_OFF3
   "Carrier_44_G120DStatusWord.6" AT %I2562.6 : Bool;   // Bit_06_LOCK_OUT
   "Carrier_44_G120DStatusWord.7" AT %I2562.7 : Bool;   // Bit_07_WARN
   "Carrier_44_G120DStatusWord.8" AT %I2563.0 : Bool;   // Bit_08_NO_DEVIATION
   "Carrier_44_G120DStatusWord.9" AT %I2563.1 : Bool;   // Bit_09_CONTR_PLC
   "Carrier_44_G120DStatusWord.10" AT %I2563.2 : Bool;   // Bit_10_F_MAX
   "Carrier_44_G120DStatusWord.11" AT %I2563.3 : Bool;   // Bit_11_LIMIT_REACHED
   "Carrier_44_G120DStatusWord.12" AT %I2563.4 : Bool;   // Bit_12_BRAKE_OPEN
   "Carrier_44_G120DStatusWord.13" AT %I2563.5 : Bool;   // Bit_13_NO_OVERTEMP
   "Carrier_44_G120DStatusWord.14" AT %I2563.6 : Bool;   // Bit_14_CW_CCW
   "Carrier_44_G120DStatusWord.15" AT %I2563.7 : Bool;   // Bit_15_OVERL
   "Carrier_44_Slot2_Input" AT %IW2564 : Word;   // SLOT 2 INPUT WORD
   "Carrier_44_CrashDetectSW" AT %I2564.0 : Bool;   // CRASH DETECT SW
   "Carrier_44_SpareSafetyInput(2_1)" AT %I2564.1 : Bool;   // SPARE SAFETY INPUT
   "Carrier_44_SpareSafetyInput(2_2)" AT %I2564.2 : Bool;   // SPARE SAFETY INPUT
   "Carrier_44_SpareSafetyInput(2_3)" AT %I2564.3 : Bool;   // SPARE SAFETY INPUT
   "Carrier_44_SpareSafetyInput(2_4)" AT %I2564.4 : Bool;   // SPARE SAFETY INPUT
   "Carrier_44_SpareSafetyInput(2_5)" AT %I2564.5 : Bool;   // SPARE SAFETY INPUT
   "Carrier_44_SpareSafetyInput(2_6)" AT %I2564.6 : Bool;   // SPARE SAFETY INPUT
   "Carrier_44_SpareSafetyInput(2_7)" AT %I2564.7 : Bool;   // SPARE SAFETY INPUT
   "Carrier_44_Slot3_SafetyOutput" AT %IW2565 : Word;   // SLOT 3 SAFETY OUTPUT WORD
   "Carrier_44_Crash_Detect_OK" AT %I2565.0 : Bool;   // CARRIER CRASH DETECT
   "Carrier_44_SpareSafetyOutput(3_1)" AT %I2565.1 : Bool;   // SPARE SAFETY OUTPUT
   "Carrier_44_SpareSafetyOutput(3_2)" AT %I2565.2 : Bool;   // SPARE SAFETY OUTPUT
   "Carrier_44_SpareSafetyOutput(3_3)" AT %I2565.3 : Bool;   // SPARE SAFETY OUTPUT
   "Carrier_44_SpareSafetyOutput(3_4)" AT %I2565.4 : Bool;   // SPARE SAFETY OUTPUT
   "Carrier_44_SpareSafetyOutput(3_5)" AT %I2565.5 : Bool;   // SPARE SAFETY OUTPUT
   "Carrier_44_SpareSafetyOutput(3_6)" AT %I2565.6 : Bool;   // SPARE SAFETY OUTPUT
   "Carrier_44_SpareSafetyOutput(3_7)" AT %I2565.7 : Bool;   // SPARE SAFETY OUTPUT
   "Carrier_44_Slot4_Input" AT %IW2566 : Word;   // SLOT 4 INPUT WORD
   "Carrier_44_480VPowerOn_MDCB1" AT %I2566.0 : Bool;   // 480 VAC POWER ON MDCB 1
   "Carrier_44_SpareInput(4_1)" AT %I2566.1 : Bool;   // SPARE INPUT
   "Carrier_44_SpareInput(4_2)" AT %I2566.2 : Bool;   // SPARE INPUT
   "Carrier_44_SitopSelectStatus" AT %I2566.3 : Bool;   // SITOP SELECT STATUS
   "Carrier_44_DCsupplyOnPSCB2" AT %I2566.4 : Bool;   // DC SUPPLY ON PSCB 2
   "Carrier_44_SpareInput(4_5)" AT %I2566.5 : Bool;   // SPARE INPUT
   "Carrier_44_SpareInput(4_6)" AT %I2566.6 : Bool;   // SPARE INPUT
   "Carrier_44_SpareInput(4_7)" AT %I2566.7 : Bool;   // SPARE INPUT
   "Carrier_44_PB1_ProdHoldLH" AT %I2567.0 : Bool;   // PB 1 PRODUCTION HOLD LH
   "Carrier_44_PB2_ResetLH" AT %I2567.1 : Bool;   // PB 2 RESET LH
   "Carrier_44_PB3_ProdHoldRH" AT %I2567.2 : Bool;   // PB 3 PRODUCTION HOLD RH
   "Carrier_44_PB4_ResetRH" AT %I2567.3 : Bool;   // PB 4 RESET RH
   "Carrier_44_SpareInput(4_14)" AT %I2567.4 : Bool;   // SPARE INPUT
   "Carrier_44_SpareInput(4_15)" AT %I2567.5 : Bool;   // SPARE INPUT
   "Carrier_44_SpareInput(4_16)" AT %I2567.6 : Bool;   // SPARE INPUT
   "Carrier_44_SpareInput(4_17)" AT %I2567.7 : Bool;   // SPARE INPUT
   "Carrier_44_Slot5_Output" AT %IW2568 : Word;   // SLOT 5 OUTPUT WORD
   "Carrier_44_IRD400_HMI_24VDC_ENABLE" AT %I2568.0 : Bool;   // IRD 400 PANEL HMI 24V DC POWER
   "Carrier_44_FaultLight_LH" AT %I2568.1 : Bool;   // FAULT LIGHT LH
   "Carrier_44_RunLight_LH" AT %I2568.2 : Bool;   // RUN LIGHT LH
   "Carrier_44_FaultLight_RH" AT %I2568.3 : Bool;   // FAULT LIGHT RH
   "Carrier_44_RunLight_RH" AT %I2568.4 : Bool;   // RUN LIGHT RH